DATA_BLOCK "T-104_Write_TO_Centrifuge_DB"   // DB309
TITLE = Signal Exchange between R-201<->Reactor_Selector
{ S7_Optimized_Access := 'TRUE' }
VERSION : 0.1
   VAR
      Wait : Bool;
      Started : Bool;   // Start Sequence
      Ready : Bool;
      Stop : Bool;   // Stop Sequence
      Abort : Bool;   // Abort Sequence
      Complete : Bool;
      Release : Bool;
      PARA : Bool;
      Initialization : Bool;
      PM : Bool;
      Monitoring : Bool;
      PumpingOut : Bool;   // Transfer to Cooling Tank
      PumpsOff : Bool;
      Held : Bool;   // Held Sequence
   END_VAR
BEGIN
END_DATA_BLOCK

DATA_BLOCK "T-104_Read_FROM_Centrifuge_DB"   // DB324
TITLE = Signal Exchange between R-201<->Reactor_Selector
{ S7_Optimized_Access := 'TRUE' }
VERSION : 0.1
   VAR
      StartTank : Bool;
      ReqWater : Bool;
      StopReqWater : Bool;
      Transfering : Bool;
      Pumps_OFF : Bool;
      Abort : Bool;
      Abort_Done : Bool;
      "Transfer_To_T-103_Done" : Bool;
      Idle : Bool;
   END_VAR
BEGIN
END_DATA_BLOCK

// folder: State MACHINE/1)Tanks/Tank T-104 (Water System)/T-104 <---> R-201

DATA_BLOCK "T-104_Write_TO_R-201_DB"   // DB287
TITLE = Signal Exchange between R-201<->Reactor_Selector
{ S7_Optimized_Access := 'TRUE' }
VERSION : 0.1
   VAR
      TankStarted : Bool;   // Start Sequence
      TankReady : Bool;
      Stop : Bool;   // Stop Sequence
      Abort : Bool;   // Abort Sequence
      PumpingOut : Bool;   // Transfer to Cooling Tank
      PumpsOff : Bool;
      Held : Bool;   // Held Sequence
   END_VAR
BEGIN
END_DATA_BLOCK

DATA_BLOCK "T-104_Read_FROM_R-201_DB"   // DB288
TITLE = Signal Exchange between R-201<->Reactor_Selector
{ S7_Optimized_Access := 'TRUE' }
VERSION : 0.1
   VAR
      StartTank : Bool;
      ReqWaterToWash : Bool;
      StopReqWaterToWash : Bool;
      ReqWater : Bool;
      StopReqWaterToPouring : Bool;
      Release : Bool;
      Abort : Bool;
      Abort_Done : Bool;
      Idle : Bool;
   END_VAR
BEGIN
END_DATA_BLOCK

// folder: State MACHINE/1)Tanks/Tank T-104 (Water System)/T-104 <---> R-202

DATA_BLOCK "T-104_Write_TO_R-202_DB"   // DB317
TITLE = Signal Exchange between R-201<->Reactor_Selector
{ S7_Optimized_Access := 'TRUE' }
VERSION : 0.1
   VAR
      TankStarted : Bool;   // Start Sequence
      TankReady : Bool;
      Stop : Bool;   // Stop Sequence
      Abort : Bool;   // Abort Sequence
      PumpingOut : Bool;   // Transfer to Cooling Tank
      PumpsOff : Bool;
      Held : Bool;   // Held Sequence
   END_VAR
BEGIN
END_DATA_BLOCK

DATA_BLOCK "T-104_Read_FROM_R-202_DB"   // DB318
TITLE = Signal Exchange between R-201<->Reactor_Selector
{ S7_Optimized_Access := 'TRUE' }
VERSION : 0.1
   VAR
      StartTank : Bool;
      ReqWaterToWash : Bool;
      StopReqWaterToWash : Bool;
      ReqWater : Bool;
      StopReqWaterToPouring : Bool;
      Release : Bool;
      Abort : Bool;
      Abort_Done : Bool;
      Idle : Bool;
   END_VAR
BEGIN
END_DATA_BLOCK

// folder: State MACHINE/1)Tanks/Tank T-104 (Water System)/T-104 <---> T-101

DATA_BLOCK "T-104_Read_FROM_T-101_DB"   // DB334
TITLE = Signal Exchange between R-201<->Reactor_Selector
{ S7_Optimized_Access := 'TRUE' }
VERSION : 0.1
   VAR
      StartTank : Bool;
      ReqWaterToWash : Bool;
      StopReqWaterToWash : Bool;
      ReqWaterToMix : Bool;
      StopReqWaterToMix : Bool;
      Release : Bool;
      Abort : Bool;
      Abort_Done : Bool;
      Idle : Bool;
   END_VAR
BEGIN
END_DATA_BLOCK

DATA_BLOCK "T-104_Write_TO_T-101_DB"   // DB341
TITLE = Signal Exchange between R-201<->Reactor_Selector
{ S7_Optimized_Access := 'TRUE' }
VERSION : 0.1
   VAR
      Wait : Bool;
      Started : Bool;   // Start Sequence
      Ready : Bool;
      Stop : Bool;   // Stop Sequence
      Abort : Bool;   // Abort Sequence
      Complete : Bool;
      Release : Bool;
      PARA : Bool;
      Initialization : Bool;
      PM : Bool;
      Monitoring : Bool;
      PumpingOut : Bool;   // Transfer to Cooling Tank
      PumpsOff : Bool;
      Held : Bool;   // Held Sequence
   END_VAR
BEGIN
END_DATA_BLOCK

// folder: State MACHINE/1)Tanks/Tank T-104 (Water System)/T-104 <---> T-102

DATA_BLOCK "T-104_Read_FROM_T-102_DB"   // DB337
TITLE = Signal Exchange between R-201<->Reactor_Selector
{ S7_Optimized_Access := 'TRUE' }
VERSION : 0.1
   VAR
      StartTank : Bool;
      ReqWaterToWash : Bool;
      StopReqWaterToWash : Bool;
      ReqWaterToMix : Bool;
      StopReqWaterToMix : Bool;
      Release : Bool;
      Abort : Bool;
      Abort_Done : Bool;
      Idle : Bool;
   END_VAR
BEGIN
END_DATA_BLOCK

DATA_BLOCK "T-104_Write_TO_T-102_DB"   // DB338
TITLE = Signal Exchange between R-201<->Reactor_Selector
{ S7_Optimized_Access := 'TRUE' }
VERSION : 0.1
   VAR
      Wait : Bool;
      Started : Bool;   // Start Sequence
      Ready : Bool;
      Stop : Bool;   // Stop Sequence
      Abort : Bool;   // Abort Sequence
      Complete : Bool;
      Release : Bool;
      PARA : Bool;
      Initialization : Bool;
      PM : Bool;
      Monitoring : Bool;
      PumpingOut : Bool;   // Transfer to Cooling Tank
      PumpsOff : Bool;
      Held : Bool;   // Held Sequence
   END_VAR
BEGIN
END_DATA_BLOCK

// folder: State MACHINE/2)Reactors/Reactor R-201

DATA_BLOCK "R-201_DB"   // DB268
{ S7_Optimized_Access := 'TRUE' }
VERSION : 0.1
   VAR
      Cmds : "UnitCmds";
      Status : Struct
         Initializing : Bool;
         Ready : Bool;
         Running : Bool;
         PouringRunning : Bool;
         TankWashRunning : Bool;
         TubeWashRunning : Bool;
         Aborting : Bool;
         Status : Int;   // 1=Idle, 2=Running, 3=Stopping, 4=Held, 5=Holding
         "Step" : Int;
         State : Int;
      END_STRUCT;
      OS : Struct
         bit : Array[0..15] of Bool;   // One Shot Bit
      END_STRUCT;
      Equipments : Struct
         Valves : Struct
            "XV-2013" : "Cmd";
            "XV-2011" : "Cmd";
            "XV-2021" : "Cmd";
            "XV-1043" : "Cmd";
            "FV-2011" : "Cmd";
            "FV-2021" : "Cmd";
         END_STRUCT;
         Pumps : Struct
            "P-201A" : "Cmd";
            "P-201B" : "Cmd";
         END_STRUCT;
         VFD : Struct
            "VFD-2011" : "Cmd";
         END_STRUCT;
      END_STRUCT;
      "Time" : Struct
         "Pre-Mix" : Time;   // Pre-Mix Time Displaying in the HMI
         pH_Delay : Time;   // pH Stabilize Time Displaying in the HMI
         Reaction : Time;   // Reaction Time Displaying in the HMI
         Wash : Time;   // Wash Time Displaying in the HMI
         Tube : Time;   // Tube Wash Time Displaying in the HMI
      END_STRUCT;
      PmpSel : Struct
         "P-201AB" : Int := 1;
      END_STRUCT;
   END_VAR
BEGIN
END_DATA_BLOCK

DATA_BLOCK "R-201_SEQ_DB"   // DB271
{ S7_Optimized_Access := 'TRUE' }
VERSION : 0.1
// stored: InstanceOfName R-201_SEQ
"R-201_SEQ"
BEGIN
END_DATA_BLOCK

DATA_BLOCK "R-201_Recipe"   // DB303
{ S7_Optimized_Access := 'TRUE' }
VERSION : 0.1
   VAR RETAIN
      Water : Real;   // Amount of Water to the Reactor before Pouring
   END_VAR
   VAR
      Temperature : Real := 80.0;   // Reactor Temperature
      MinLevelMixerOn : Real := 19.0;   // Minimum Level to Run the Mixer
      X_Flow : Real := 1.0;   // T-101(X) Flow to Transfer to Reactor
      Y_Flow : Real := 1.5;   // T-102(Y) Flow to Transfer to Reactor with pH Stability.
      X_Volume : Real;   // T-101(X) Volume to Transfer to Reactor
      LastWaterVolume : Real := 120.0;
      pH : Real := 8.0;   // pH Setpoint to the Reactor
      "Pre-Mix_Time" : Time := T#5m;   // Pre-Mix Time to the T-101 and T-102 before Transfer to Reactor
      pHStab_Time : Time := T#1m;   // Time to Stabilize the pH
      Reaction_Time : Time := T#22.5h;   // Reaction Time
   END_VAR
BEGIN
END_DATA_BLOCK

DATA_BLOCK "R-201_Aux_DB"   // DB354
{ S7_Optimized_Access := 'TRUE' }
VERSION : 0.1
   VAR
      "Real" : Struct
         "HFC-201" : Struct   // Heater
            SP : Real;
            Min : Real;   // Heater Minimum Temperature
            Max : Real;   // Heater Maximum Temperature
         END_STRUCT;
         PH : Struct   // pH Controller
            SP : Real;   // pH Set Point
            Min : Real;
            Max : Real;
         END_STRUCT;
         "FIC-2011" : Struct   // Fow Controller
            SP : Real := 1.0;   // Flow Setpoint
         END_STRUCT;
         "FIC-2021" : Struct
            SP : Real := 1.5;   // Flow Setpoint
         END_STRUCT;
         "T-101" : Struct
            TOTVolSP : Real;
         END_STRUCT;
         "LT-2011" : Struct
            Min : Real;
         END_STRUCT;
         "FT-1043" : Struct
            SP : Real;
         END_STRUCT;
         "VFD-R201" : Struct
            Start : Bool;
            Stop : Bool;
         END_STRUCT;
      END_STRUCT;
      "Timer" : Struct
         PreMix : IEC_TIMER;   // Timer Premix
         StabpH : IEC_TIMER;
         Reactor : IEC_TIMER;
         FlushOut : IEC_TIMER;
         MixToClean : IEC_TIMER;
         "XV-2013" : IEC_TIMER;
         "XV-2011" : IEC_TIMER;
         "XV-2021" : IEC_TIMER;
         "XV-1043" : IEC_TIMER;
         "FV-2011" : IEC_TIMER;
         "FV-2021" : IEC_TIMER;
      END_STRUCT;
      "Bool" : Struct
         PreMixT_En : Bool;   // Pre-Mix Timer Enable
         PreMixT_Reset : Bool;
         StabpHTEnStep : Bool;   // Stabilizer Timer Enable
         StabpHTEn : Bool;
         StabpHTEn_Reset : Bool;
         ReactorTEn : Bool;   // Enable Reacting time for the Reactor
         ReactorT_Reset : Bool;
         FlushOutTEn : Bool;
         MixToCleanTEn : Bool;   // Enable Timer to clean the reactor after Reacting
         MixToCleanT_Reset : Bool;
         TOff : Bool;   // Turning Off Valves
         Transitions : Struct
            TankEmpty : Bool;
         END_STRUCT;
      END_STRUCT;
      Constants : Struct
         CmdDelay : Time := T#2s;
      END_STRUCT;
   END_VAR
BEGIN
   "Timer".FlushOut.PT := T#5S;
   "Timer".PreMix.PT := T#5m;
   "Timer".StabpH.PT := T#1m;
   "Timer".MixToClean.PT := T#10M;
   "Timer".Reactor.PT := T#22.5h;
END_DATA_BLOCK

DATA_BLOCK "R-201_HMI_DB"   // DB358
{ S7_Optimized_Access := 'TRUE' }
VERSION : 0.1
   VAR
      FromHMI : "FromHMI";
      ToHMI : "ToHMI";
   END_VAR
BEGIN
END_DATA_BLOCK

// folder: State MACHINE/2)Reactors/Reactor R-201/Control R-201

DATA_BLOCK "R-201_Control_SEQ_DB"   // DB283
{ S7_Optimized_Access := 'TRUE' }
VERSION : 0.1
// stored: InstanceOfName R-201_Control
"R-201_Control"
BEGIN
END_DATA_BLOCK

DATA_BLOCK "R-201_Control_DB"   // DB300
{ S7_Optimized_Access := 'TRUE' }
VERSION : 0.1
   VAR
      FromHMI : Struct
         Start : Bool;
         Initialize : Bool;
         TankWash : Bool;
         TubeWash : Bool;
         Abort : Bool;
      END_STRUCT;
      Cmds : Struct
         Start : Bool;
         Initialize : Bool;
         TankWash : Bool;
         TubeWash : Bool;
         TransferToCoolingTank : Bool;
         Abort : Bool;
      END_STRUCT;
      Status : Struct
         Starting : Bool;
         Aborting : Bool;
      END_STRUCT;
      OS : Struct
         bit : Array[0..15] of Bool;   // One Shot Bit
      END_STRUCT;
   END_VAR
BEGIN
END_DATA_BLOCK

// folder: State MACHINE/2)Reactors/Reactor R-201/Control R-201/Control <---> R-201

DATA_BLOCK "Control_Write_TO_R-201_DB"   // DB277
TITLE = Signal Exchange between R-201<->Reactor_Selector
{ S7_Optimized_Access := 'TRUE' }
VERSION : 0.1
   VAR
      Wait : Bool;
      Start : Bool;   // Start Sequence
      Stop : Bool;   // Stop Sequence
      Abort : Bool;   // Abort Sequence
      Complete : Bool;
      Release : Bool;
      PARA : Bool;
      Initialization : Bool;
      PM : Bool;
      Running : Bool;
      WaitForTransfer : Bool;
      "Transfer_To_T-103" : Bool;   // Transfer to Cooling Tank
      TankWash : Bool;
      TubingWash : Bool;
      Held : Bool;   // Held Sequence
   END_VAR
BEGIN
END_DATA_BLOCK

DATA_BLOCK "Control_Read_FROM_R-201_DB"   // DB280
TITLE = Signal Exchange between R-201<->Reactor_Selector
{ S7_Optimized_Access := 'TRUE' }
VERSION : 0.1
   VAR
      ReactorStarted : Bool;
      Initialization_Done : Bool;
      Reacting_Done : Bool;
      Abort_Done : Bool;
      "Transfer_To_T-103_Done" : Bool;
      TankWash_done : Bool;
      TubeWash_Done : Bool;
      Idle : Bool;
   END_VAR
BEGIN
END_DATA_BLOCK

// folder: State MACHINE/2)Reactors/Reactor R-201/R-201 <---> Control

DATA_BLOCK "R-201_Write_TO_Control_DB"   // DB281
TITLE = Signal Exchange between R-201<->Reactor_Selector
{ S7_Optimized_Access := 'TRUE' }
VERSION : 0.1
   VAR
      ReactorStarted : Bool;
      Initialization_Done : Bool;
      Reacting_Done : Bool;
      Abort_Done : Bool;
      "Transfer_To_T-103_Done" : Bool;
      TankWash_done : Bool;
      TubeWash_Done : Bool;
      Idle : Bool;
   END_VAR
BEGIN
END_DATA_BLOCK

DATA_BLOCK "R-201_Read_FROM_Control_DB"   // DB282
TITLE = Signal Exchange between R-201<->Reactor_Selector
{ S7_Optimized_Access := 'TRUE' }
VERSION : 0.1
   VAR
      Wait : Bool;
      Start : Bool;   // Start Sequence
      Stop : Bool;   // Stop Sequence
      Abort : Bool;   // Abort Sequence
      Complete : Bool;
      Release : Bool;
      PARA : Bool;
      Initialization : Bool;
      PM : Bool;
      Running : Bool;
      WaitForTransfer : Bool;
      "Transfer_To_T-103" : Bool;   // Transfer to Cooling Tank
      TankWash : Bool;
      TubingWash : Bool;
      Held : Bool;   // Held Sequence
   END_VAR
BEGIN
END_DATA_BLOCK

// folder: State MACHINE/2)Reactors/Reactor R-201/R-201 <---> T-101

DATA_BLOCK "R-201_Read_FROM_T-101_DB"   // DB307
TITLE = Signal Exchange between R-201<->Reactor_Selector
{ S7_Optimized_Access := 'TRUE' }
VERSION : 0.1
   VAR
      TankStarted : Bool;   // Start Sequence
      Recirculating : Bool;
      PupmsOFF : Bool;   // Stop Sequence
      Abort : Bool;   // Abort Sequence
      RouteOpened : Bool;   // Transfer to Cooling Tank
      Idle : Bool;   // Held Sequence
   END_VAR
BEGIN
END_DATA_BLOCK

DATA_BLOCK "R-201_Write_TO_T-101_DB"   // DB327
TITLE = Signal Exchange between R-201<->Reactor_Selector
{ S7_Optimized_Access := 'TRUE' }
VERSION : 0.1
   VAR
      StartPouring : Bool;
      ReactorStarted : Bool;
      OpenRoute : Bool;
      RouteOpened : Bool;
      Transfering : Bool;
      FillingDone : Bool;
      Abort : Bool;
      Abort_Done : Bool;
      ReleaseTank : Bool;
      Idle : Bool;
   END_VAR
BEGIN
END_DATA_BLOCK

// folder: State MACHINE/2)Reactors/Reactor R-201/R-201 <---> T-102

DATA_BLOCK "R-201_Read_FROM_T-102_DB"   // DB316
TITLE = Signal Exchange between R-201<->Reactor_Selector
{ S7_Optimized_Access := 'TRUE' }
VERSION : 0.1
   VAR
      TankStarted : Bool;   // Start Sequence
      Recirculating : Bool;
      PupmsOFF : Bool;   // Stop Sequence
      Abort : Bool;   // Abort Sequence
      RouteOpened : Bool;   // Transfer to Cooling Tank
      Idle : Bool;   // Held Sequence
   END_VAR
BEGIN
END_DATA_BLOCK

DATA_BLOCK "R-201_Write_TO_T-102_DB"   // DB319
TITLE = Signal Exchange between R-201<->Reactor_Selector
{ S7_Optimized_Access := 'TRUE' }
VERSION : 0.1
   VAR
      StartPouring : Bool;
      ReactorStarted : Bool;
      OpenRoute : Bool;
      RouteOpened : Bool;
      Transfering : Bool;
      FillingDone : Bool;
      Abort : Bool;
      Abort_Done : Bool;
      ReleaseTank : Bool;
      Idle : Bool;
   END_VAR
BEGIN
END_DATA_BLOCK

// folder: State MACHINE/2)Reactors/Reactor R-201/R-201 <---> T-103 (CoolingTank)

DATA_BLOCK "R-201_Write_TO_T-103_DB"   // DB293
TITLE = Signal Exchange between R-201<->Reactor_Selector
{ S7_Optimized_Access := 'TRUE' }
VERSION : 0.1
   VAR
      StartTank : Bool;
      OpenRoute : Bool;
      Transfering : Bool;
      TubWash_Done : Bool;
      Abort : Bool;
      Abort_Done : Bool;
      "Transfer_To_T-103_Done" : Bool;
      Idle : Bool;
   END_VAR
BEGIN
END_DATA_BLOCK

DATA_BLOCK "R-201_Read_FROM_T-103_DB"   // DB296
TITLE = Signal Exchange between R-201<->Reactor_Selector
{ S7_Optimized_Access := 'TRUE' }
VERSION : 0.1
   VAR
      TankStarted : Bool;   // Start Sequence
      Stop : Bool;   // Stop Sequence
      Abort : Bool;   // Abort Sequence
      RouteOpened : Bool;   // Transfer to Cooling Tank
      Release : Bool;
      Held : Bool;   // Held Sequence
   END_VAR
BEGIN
END_DATA_BLOCK

// folder: State MACHINE/2)Reactors/Reactor R-201/R-201 <---> T-104 (WaterSystem)

DATA_BLOCK "R-201_Write_TO_T-104_DB"   // DB294
TITLE = Signal Exchange between R-201<->Reactor_Selector
{ S7_Optimized_Access := 'TRUE' }
VERSION : 0.1
   VAR
      StartTank : Bool;
      ReqWaterToWash : Bool;
      StopReqWaterToWash : Bool;
      ReqWater : Bool;
      StopReqWaterToPouring : Bool;
      Release : Bool;
      Abort : Bool;
      Abort_Done : Bool;
      Idle : Bool;
   END_VAR
BEGIN
END_DATA_BLOCK

DATA_BLOCK "R-201_Read_FROM_T-104_DB"   // DB295
TITLE = Signal Exchange between R-201<->Reactor_Selector
{ S7_Optimized_Access := 'TRUE' }
VERSION : 0.1
   VAR
      Wait : Bool;
      TankStarted : Bool;   // Start Sequence
      Ready : Bool;
      Stop : Bool;   // Stop Sequence
      Abort : Bool;   // Abort Sequence
      PumpingOut : Bool;   // Transfer to Cooling Tank
      PumpsOff : Bool;
      Held : Bool;   // Held Sequence
   END_VAR
BEGIN
END_DATA_BLOCK

// folder: State MACHINE/2)Reactors/Reactor R-202

DATA_BLOCK "R-202_DB"   // DB269
{ S7_Optimized_Access := 'TRUE' }
VERSION : 0.1
   VAR
      FromHMI : Struct
         Start : Bool;
         Initialize : Bool;
         TankWash : Bool;
         TubeWash : Bool;
         TransferToCoolingTank : Bool;
         Abort : Bool;
      END_STRUCT;
      Cmds : "UnitCmds";
      Status : Struct
         Initializing : Bool;
         Ready : Bool;
         Running : Bool;
         PouringRunning : Bool;
         TankWashRunning : Bool;
         TubeWashRunning : Bool;
         Aborting : Bool;
         Status : Int;   // 1=Idle, 2=Running, 3=Stopping, 4=Held, 5=Holding
         "Step" : Int;
         State : Int;
      END_STRUCT;
      OS : Struct
         bit : Array[0..15] of Bool;   // One Shot Bit
      END_STRUCT;
      Equipments : Struct
         Valves : Struct
            "XV-2023" : "Cmd";
            "XV-2012" : "Cmd";
            "XV-2022" : "Cmd";
            "XV-1044" : "Cmd";
            "FV-2012" : "Cmd";
            "FV-2022" : "Cmd";
         END_STRUCT;
         Pumps : Struct
            "P-202A" : "Cmd";
            "P-202B" : "Cmd";
         END_STRUCT;
         VFD : Struct
            "VFD-2021" : "Cmd";
         END_STRUCT;
      END_STRUCT;
      "Time" : Struct
         "Pre-Mix" : Time;   // Pre-Mix Time Displaying in the HMI
         PH_Delay : Time;   // pH Stabilize Time Displaying in the HMI
         Reaction : Time;   // Reaction Time Displaying in the HMI
         Wash : Time;   // Wash Time Displaying in the HMI
         Tube : Time;   // Tube Wash Time Displaying in the HMI
      END_STRUCT;
      PmpSel : Struct
         "P-202AB" : Int := 1;
      END_STRUCT;
   END_VAR
BEGIN
END_DATA_BLOCK

DATA_BLOCK "R-202_SEQ_DB"   // DB286
{ S7_Optimized_Access := 'TRUE' }
VERSION : 0.1
// stored: InstanceOfName R-202_SEQ
"R-202_SEQ"
BEGIN
END_DATA_BLOCK

DATA_BLOCK "R-202_Recipe"   // DB304
{ S7_Optimized_Access := 'TRUE' }
VERSION : 0.1
   VAR RETAIN
      Water : Real;   // Amount of Water to the Reactor before Pouring
   END_VAR
   VAR
      Temperature : Real := 80.0;   // Reactor Temperature
      MinLevelMixerOn : Real := 19.0;   // Minimum Level to Run the Mixer
      X_Flow : Real := 1.0;   // T-101(X) Flow to Transfer to Reactor
      Y_Flow : Real := 1.5;   // T-102(Y) Flow to Transfer to Reactor with pH Stability.
      X_Volume : Real;   // T-101(X) Volume to Transfer to Reactor
      LastWaterVolume : Real := 120.0;
      pH : Real := 8.0;   // pH Setpoint to the Reactor
      "Pre-Mix_Time" : Time := T#5m;   // Pre-Mix Time to the T-101 and T-102 before Transfer to Reactor
      pHStab_Time : Time := T#1m;   // Time to Stabilize the pH
      Reaction_Time : Time := T#22.5h;   // Reaction Time
   END_VAR
BEGIN
END_DATA_BLOCK

DATA_BLOCK "R-202_Aux_DB"   // DB365
{ S7_Optimized_Access := 'TRUE' }
VERSION : 0.1
   VAR
      "Real" : Struct
         "HFC-201" : Struct   // Heater
            SP : Real;
            Min : Real;   // Heater Minimum Temperature
            Max : Real;   // Heater Maximum Temperature
         END_STRUCT;
         PH : Struct   // pH Controller
            SP : Real;   // pH Set Point
            Min : Real;
            Max : Real;
         END_STRUCT;
         "FIC-2012" : Struct   // Fow Controller
            SP : Real;   // Flow Setpoint
         END_STRUCT;
         "FIC-2022" : Struct
            SP : Real := 1.0;   // Flow Setpoint
         END_STRUCT;
         "T-101" : Struct
            TOTVolSP : Real;
         END_STRUCT;
         "LT-2021" : Struct
            Min : Real;
         END_STRUCT;
         "FT-1044" : Struct
            SP : Real;
         END_STRUCT;
         "VFD-R202" : Struct
            Start : Bool;
            Stop : Bool;
         END_STRUCT;
      END_STRUCT;
      "Timer" : Struct
         PreMix : IEC_TIMER;   // Timer Premix
         StabpH : IEC_TIMER;
         Reactor : IEC_TIMER;
         FlushOut : IEC_TIMER;
         MixToClean : IEC_TIMER;
         "XV-2023" : IEC_TIMER;
         "XV-2012" : IEC_TIMER;
         "XV-2022" : IEC_TIMER;
         "XV-1044" : IEC_TIMER;
         "FV-2012" : IEC_TIMER;
         "FV-2022" : IEC_TIMER;
      END_STRUCT;
      "Bool" : Struct
         PreMixT_En : Bool;   // Pre-Mix Timer Enable
         PreMixT_Reset : Bool;
         StabpHTEnStep : Bool;   // Stabilizer Timer Enable
         StabpHTEn : Bool;   // Stabilizer Timer Enable
         StabpHTEn_Reset : Bool;
         ReactorTEn : Bool;   // Enable Reacting time for the Reactor
         ReactorT_Reset : Bool;
         FlushOutTEn : Bool;
         MixToCleanTEn : Bool;   // Enable Timer to clean the reactor after Reacting
         MixToCleanT_Reset : Bool;
         TOff : Bool;   // Turning Off Valves
         Transitions : Struct
            TankEmpty : Bool;
         END_STRUCT;
      END_STRUCT;
      Constants : Struct
         CmdDelay : Time := T#2s;
      END_STRUCT;
   END_VAR
BEGIN
   "Timer".FlushOut.PT := T#5S;
   "Timer".PreMix.PT := T#5m;
   "Timer".StabpH.PT := T#1m;
   "Timer".MixToClean.PT := T#10M;
   "Timer".Reactor.PT := T#21.5h;
END_DATA_BLOCK

DATA_BLOCK "R-202_HMI_DB"   // DB367
{ S7_Optimized_Access := 'TRUE' }
VERSION : 0.1
   VAR
      FromHMI : "FromHMI";
      ToHMI : "ToHMI";
   END_VAR
BEGIN
END_DATA_BLOCK

// folder: State MACHINE/2)Reactors/Reactor R-202/Control R-202

DATA_BLOCK "R-202_Control_SEQ_DB"   // DB290
{ S7_Optimized_Access := 'TRUE' }
VERSION : 0.1
// stored: InstanceOfName R-202_Control
"R-202_Control"
BEGIN
END_DATA_BLOCK

DATA_BLOCK "R-202_Control_DB"   // DB344
{ S7_Optimized_Access := 'TRUE' }
VERSION : 0.1
   VAR
      FromHMI : Struct
         Start : Bool;
         Initialize : Bool;
         TankWash : Bool;
         TubeWash : Bool;
         Abort : Bool;
      END_STRUCT;
      Cmds : Struct
         Start : Bool;
         Initialize : Bool;
         TankWash : Bool;
         TubeWash : Bool;
         Abort : Bool;
      END_STRUCT;
      Status : Struct
         Starting : Bool;
         Aborting : Bool;
      END_STRUCT;
      OS : Struct
         bit : Array[0..15] of Bool;   // One Shot Bit
      END_STRUCT;
   END_VAR
BEGIN
END_DATA_BLOCK

// folder: State MACHINE/2)Reactors/Reactor R-202/Control R-202/Control <---> R-202

DATA_BLOCK "Control_Write_TO_R-202_DB"   // DB270
TITLE = Signal Exchange between R-201<->Reactor_Selector
{ S7_Optimized_Access := 'TRUE' }
VERSION : 0.1
   VAR
      Wait : Bool;
      Start : Bool;   // Start Sequence
      Stop : Bool;   // Stop Sequence
      Abort : Bool;   // Abort Sequence
      Complete : Bool;
      Release : Bool;
      PARA : Bool;
      Initialization : Bool;
      PM : Bool;
      Running : Bool;
      "Transfer_To_T-103" : Bool;   // Transfer to Cooling Tank
      TankWash : Bool;
      TubingWash : Bool;
      Held : Bool;   // Held Sequence
   END_VAR
BEGIN
END_DATA_BLOCK

DATA_BLOCK "Control_Read_FROM_R-202_DB"   // DB273
TITLE = Signal Exchange between R-201<->Reactor_Selector
{ S7_Optimized_Access := 'TRUE' }
VERSION : 0.1
   VAR
      ReactorStarted : Bool;
      Initialization_Done : Bool;
      Reacting_Done : Bool;
      Abort_Done : Bool;
      "Transfer_To_T-103_Done" : Bool;
      TankWash_done : Bool;
      TubeWash_Done : Bool;
      Idle : Bool;
   END_VAR
BEGIN
END_DATA_BLOCK

// folder: State MACHINE/2)Reactors/Reactor R-202/R-202 <---> Control

DATA_BLOCK "R-202_Write_TO_Control_DB"   // DB285
TITLE = Signal Exchange between R-201<->Reactor_Selector
{ S7_Optimized_Access := 'TRUE' }
VERSION : 0.1
   VAR
      ReactorStarted : Bool;
      Initialization_Done : Bool;
      Reacting_Done : Bool;
      Abort_Done : Bool;
      "Transfer_To_T-103_Done" : Bool;
      TankWash_done : Bool;
      TubeWash_Done : Bool;
      Idle : Bool;
   END_VAR
BEGIN
END_DATA_BLOCK

DATA_BLOCK "R-202_Read_FROM_Control_DB"   // DB289
TITLE = Signal Exchange between R-201<->Reactor_Selector
{ S7_Optimized_Access := 'TRUE' }
VERSION : 0.1
   VAR
      Wait : Bool;
      Start : Bool;   // Start Sequence
      Stop : Bool;   // Stop Sequence
      Abort : Bool;   // Abort Sequence
      Complete : Bool;
      Release : Bool;
      PARA : Bool;
      Initialization : Bool;
      PM : Bool;
      Running : Bool;
      "Transfer_To_T-103" : Bool;   // Transfer to Cooling Tank
      TankWash : Bool;
      TubingWash : Bool;
      Held : Bool;   // Held Sequence
   END_VAR
BEGIN
END_DATA_BLOCK

// folder: State MACHINE/2)Reactors/Reactor R-202/R-202 <---> T-101

DATA_BLOCK "R-202_Read_FROM_T-101_DB"   // DB312
TITLE = Signal Exchange between R-201<->Reactor_Selector
{ S7_Optimized_Access := 'TRUE' }
VERSION : 0.1
   VAR
      TankStarted : Bool;   // Start Sequence
      Recirculating : Bool;
      PupmsOFF : Bool;   // Stop Sequence
      Abort : Bool;   // Abort Sequence
      RouteOpened : Bool;   // Transfer to Cooling Tank
      Idle : Bool;   // Held Sequence
   END_VAR
BEGIN
END_DATA_BLOCK

DATA_BLOCK "R-202_Write_TO_T-101_DB"   // DB329
TITLE = Signal Exchange between R-201<->Reactor_Selector
{ S7_Optimized_Access := 'TRUE' }
VERSION : 0.1
   VAR
      StartPouring : Bool;
      ReactorStarted : Bool;
      OpenRoute : Bool;
      RouteOpened : Bool;
      Transfering : Bool;
      FillingDone : Bool;
      Abort : Bool;
      Abort_Done : Bool;
      ReleaseTank : Bool;
      Idle : Bool;
   END_VAR
BEGIN
END_DATA_BLOCK

// folder: State MACHINE/2)Reactors/Reactor R-202/R-202 <---> T-102

DATA_BLOCK "R-202_Read_FROM_T-102_DB"   // DB313
TITLE = Signal Exchange between R-201<->Reactor_Selector
{ S7_Optimized_Access := 'TRUE' }
VERSION : 0.1
   VAR
      TankStarted : Bool;   // Start Sequence
      Recirculating : Bool;
      PupmsOFF : Bool;   // Stop Sequence
      Abort : Bool;   // Abort Sequence
      RouteOpened : Bool;   // Transfer to Cooling Tank
      Idle : Bool;   // Held Sequence
   END_VAR
BEGIN
END_DATA_BLOCK

DATA_BLOCK "R-202_Write_TO_T-102_DB"   // DB330
TITLE = Signal Exchange between R-201<->Reactor_Selector
{ S7_Optimized_Access := 'TRUE' }
VERSION : 0.1
   VAR
      StartPouring : Bool;
      ReactorStarted : Bool;
      OpenRoute : Bool;
      RouteOpened : Bool;
      Transfering : Bool;
      FillingDone : Bool;
      Abort : Bool;
      Abort_Done : Bool;
      ReleaseTank : Bool;
      Idle : Bool;
   END_VAR
BEGIN
END_DATA_BLOCK

// folder: State MACHINE/2)Reactors/Reactor R-202/R-202 <---> T-103 (CoolingTank)

DATA_BLOCK "R-202_Write_TO_T-103_DB"   // DB332
TITLE = Signal Exchange between R-201<->Reactor_Selector
{ S7_Optimized_Access := 'TRUE' }
VERSION : 0.1
   VAR
      StartTank : Bool;
      OpenRoute : Bool;
      Transfering : Bool;
      TubWash_Done : Bool;
      Abort : Bool;
      Abort_Done : Bool;
      "Transfer_To_T-103_Done" : Bool;
      Idle : Bool;
   END_VAR
BEGIN
END_DATA_BLOCK

DATA_BLOCK "R-202_Read_FROM_T-103_DB"   // DB343
TITLE = Signal Exchange between R-201<->Reactor_Selector
{ S7_Optimized_Access := 'TRUE' }
VERSION : 0.1
   VAR
      TankStarted : Bool;   // Start Sequence
      Stop : Bool;   // Stop Sequence
      Abort : Bool;   // Abort Sequence
      RouteOpened : Bool;   // Transfer to Cooling Tank
      Release : Bool;
      Held : Bool;   // Held Sequence
   END_VAR
BEGIN
END_DATA_BLOCK

// folder: State MACHINE/2)Reactors/Reactor R-202/R-202 <---> T-104 (WaterSystem)

DATA_BLOCK "R-202_Write_TO_T-104_DB"   // DB335
TITLE = Signal Exchange between R-201<->Reactor_Selector
{ S7_Optimized_Access := 'TRUE' }
VERSION : 0.1
   VAR
      StartTank : Bool;
      ReqWaterToWash : Bool;
      StopReqWaterToWash : Bool;
      ReqWater : Bool;
      StopReqWaterToPouring : Bool;
      Release : Bool;
      Abort : Bool;
      Abort_Done : Bool;
      Idle : Bool;
   END_VAR
BEGIN
END_DATA_BLOCK

DATA_BLOCK "R-202_Read_FROM_T-104_DB"   // DB339
TITLE = Signal Exchange between R-201<->Reactor_Selector
{ S7_Optimized_Access := 'TRUE' }
VERSION : 0.1
   VAR
      Wait : Bool;
      TankStarted : Bool;   // Start Sequence
      Ready : Bool;
      Stop : Bool;   // Stop Sequence
      Abort : Bool;   // Abort Sequence
      PumpingOut : Bool;   // Transfer to Cooling Tank
      PumpsOff : Bool;
      Held : Bool;   // Held Sequence
   END_VAR
BEGIN
END_DATA_BLOCK

// folder: State MACHINE/3)Centrifuge

DATA_BLOCK "Centrifuge_DB"   // DB266
{ S7_Optimized_Access := 'TRUE' }
VERSION : 0.1
   VAR
      Transitions : Struct
         "T-103_Empty" : Bool;
         WaterDone : Bool;
         InitialsDone : Bool;
         ReadytoRun : Bool;
         BasketFull : Bool;
      END_STRUCT;
      Timers : Struct
         BucketTimerDelay : IEC_TIMER;
      END_STRUCT;
      Cmds : "UnitCmds";
      Status : Struct
         Initializing : Bool;
         Ready : Bool;
         Running : Bool;
         PouringRunning : Bool;
         TankWashRunning : Bool;
         TubeWashRunning : Bool;
         Aborting : Bool;
         Status : Int;   // 1=Idle, 2=Running, 3=Stopping, 4=Held, 5=Holding
         "Step" : Int;
         State : Int;
      END_STRUCT;
      OS : Struct
         bit : Array[0..15] of Bool;   // One Shot Bit
      END_STRUCT;
      Equipments : Struct
         Valves : Struct
            "XV-1045" : "Cmd";
            "XV-3013" : "Cmd";
            "XV-3012" : "Cmd";
            "XV-3011" : "Cmd";
            "FV-3011" : "Cmd";
         END_STRUCT;
         Pumps : Struct
            "P-301A" : "Cmd";
            "P-301B" : "Cmd";
         END_STRUCT;
         VFD : Struct
            "C-3011" : "Centrifuge";
         END_STRUCT;
      END_STRUCT;
      "Time" : Struct
         DrySpin : Time;
      END_STRUCT;
      PmpSel : Struct   // PumpSelection
         "P-301AB" : Int := 1;   // 1=P-301A, 2=P-301B
      END_STRUCT;
   END_VAR
BEGIN
END_DATA_BLOCK

DATA_BLOCK "Centrifuge_SEQ_DB"   // DB299
{ S7_Optimized_Access := 'TRUE' }
VERSION : 0.1
// stored: InstanceOfName Centrifuge_SEQ
"Centrifuge_SEQ"
BEGIN
END_DATA_BLOCK

DATA_BLOCK "Centrifuge_Aux_DB"   // DB356
{ S7_Optimized_Access := 'TRUE' }
VERSION : 0.1
   VAR
      "Real" : Struct
         "FIC-3011" : Struct
            SP : Real := 10.0;
         END_STRUCT;
         "VFD-3011" : Struct
            SP : Real := 50.0;
         END_STRUCT;
         "FT-3011" : Struct
            SP : Real := 280.0;
         END_STRUCT;
         DryTime : Struct
            SP : Time := T#10M;
         END_STRUCT;
      END_STRUCT;
      "Int" : Struct
         CentrifugeSpeedFbk : Int;
      END_STRUCT;
      "Timer" : Struct
         "XV-1045" : IEC_TIMER;
         "XV-3013" : IEC_TIMER;
         "XV-3012" : IEC_TIMER;
         "XV-3011" : IEC_TIMER;
         "FV-3011" : IEC_TIMER;
         WaitForBucket : IEC_TIMER;
         DryingWetCake : IEC_TIMER;
         DrySpinDnDelay : IEC_TIMER;   // Dry Spin Done Delay to Finish
      END_STRUCT;
      "Bool" : Struct
         TOff : Bool;   // Turning Off Valves
         WaitForBucketEn : Bool;   // Wait for get some Level in the Bucket before Start Pumps
         DryingWetCakeEn : Bool;   // Run the Pumps after Turn off the Water to dry the wet cake
         DryingWetCake_Reset : Bool;
         DrySpinDnDelay_Enab : Bool;
         Centrifuge : Struct
            Status : Struct
               MotorRunning : Bool;
               VibrationFault : Bool;
               ESTOP : Bool;
               SystemFault : Bool;
               BasketFull : Bool;
               CoverLocked : Bool;
               FeelerRetracted : Bool;
               FeelerEngaged : Bool;
            END_STRUCT;
            Command : Struct
               Start : Bool;
               Stop : Bool;
               ESTOP : Bool := TRUE;   // ESTOP to Centrifuge, 1=OK
               RetFeelerAndReset : Bool;
               FeelerEngage : Bool;
            END_STRUCT;
         END_STRUCT;
      END_STRUCT;
      Constants : Struct
         CmdDelay : Time := T#2s;
      END_STRUCT;
   END_VAR
BEGIN
   "Timer".DryingWetCake.PT := t#30m;
   "Timer".DrySpinDnDelay.PT := T#30s;
END_DATA_BLOCK

DATA_BLOCK "Centrifuge_HMI_DB"   // DB363
{ S7_Optimized_Access := 'TRUE' }
VERSION : 0.1
   VAR
      FromHMI : "FromHMI";
      ToHMI : "ToHMI";
      FromHMI_Aux : Struct
         Start : Bool;   // Start Centrifuge
         Stop : Bool;   // Stop Centrifuge
         FeelerRetReset : Bool;   // Feeler Retrac and Reset
         FeelerEngage : Bool;   // Feeler Engage
      END_STRUCT;
   END_VAR
BEGIN
END_DATA_BLOCK

// folder: State MACHINE/3)Centrifuge/Centrifuge <---> T-103

DATA_BLOCK "Centrifuge_Write_TO_T-103_DB"   // DB310
TITLE = Signal Exchange between R-201<->Reactor_Selector
{ S7_Optimized_Access := 'TRUE' }
VERSION : 0.1
   VAR
      RequestProduct : Bool;   // Request Product
      OpenRoute : Bool;
      RouteOpened : Bool;   // Abort Sequence
      "T-103_Empty" : Bool;   // T-103 Tank empty
      BasketFull : Bool;   // Basket Full Signal
      FeelerRet : Bool;   // Feeler Retracted
      CloseRoute : Bool;
      Release : Bool;
   END_VAR
BEGIN
END_DATA_BLOCK

DATA_BLOCK "Centrifuge_Read_FROM_T-103_DB"   // DB320
TITLE = Signal Exchange between R-201<->Reactor_Selector
{ S7_Optimized_Access := 'TRUE' }
VERSION : 0.1
   VAR
      ReadyToTransfer : Bool;
      Done : Bool;
      RouteOpened : Bool;
      Transfering : Bool;
      Pumps_OFF : Bool;
      Abort : Bool;
      Abort_Done : Bool;
      "Transfer_To_T-103_Done" : Bool;
      Idle : Bool;
   END_VAR
BEGIN
END_DATA_BLOCK

// folder: State MACHINE/3)Centrifuge/Centrifuge <---> T-104

DATA_BLOCK "Centrifuge_Write_TO_T-104_DB"   // DB315
TITLE = Signal Exchange between R-201<->Reactor_Selector
{ S7_Optimized_Access := 'TRUE' }
VERSION : 0.1
   VAR
      StartTank : Bool;   // Start Sequence
      ReqWater : Bool;
      StopReqWater : Bool;
      Abort : Bool;   // Abort Sequence
      Complete : Bool;
      Release : Bool;
      PARA : Bool;
      Initialization : Bool;
      PM : Bool;
      Monitoring : Bool;
      RouteOpened : Bool;   // Transfer to Cooling Tank
      Held : Bool;   // Held Sequence
   END_VAR
BEGIN
END_DATA_BLOCK

DATA_BLOCK "Centrifuge_Read_FROM_T-104_DB"   // DB323
TITLE = Signal Exchange between R-201<->Reactor_Selector
{ S7_Optimized_Access := 'TRUE' }
VERSION : 0.1
   VAR
      Wait : Bool;
      Started : Bool;   // Start Sequence
      Ready : Bool;
      Stop : Bool;   // Stop Sequence
      Abort : Bool;   // Abort Sequence
      Complete : Bool;
      Release : Bool;
      PARA : Bool;
      Initialization : Bool;
      PM : Bool;
      Monitoring : Bool;
      PumpingOut : Bool;   // Transfer to Cooling Tank
      PumpsOff : Bool;
      Held : Bool;   // Held Sequence
   END_VAR
BEGIN
END_DATA_BLOCK

// folder: State MACHINE/4)Calcination

DATA_BLOCK "R401_TempMon_DB"   // DB20
{ S7_Optimized_Access := 'TRUE' }
AUTHOR : JLopez
VERSION : 0.1
// stored: InstanceOfName AI Monitor
"AI Monitor"
BEGIN
END_DATA_BLOCK

DATA_BLOCK "Calcination_DB"   // DB91
{ S7_Optimized_Access := 'TRUE' }
VERSION : 0.1
   VAR
      Alarms : Struct
         Communication : Struct
            Fault : Bool;
         END_STRUCT;
      END_STRUCT;
      Shutdowns : Struct
         "1 Activated" : Bool;
         "2 Activated" : Bool;
      END_STRUCT;
      MonBlockData : Struct
         Input : Struct
            AvgSP : Real;   // Average SP Furnace Temperature
            "Min Range" : Real;   // Minimum Furnace Temperature Range
            "Max Range" : Real;   // Maximun Furnace Temperature Range
            MinAvgValue : Real := 0.0;   // Min Average Hysteresis Range
            MaxAvgValue : Real := 0.0;   // Max Average Hysteresis Range
            EnableDeviationMon : Bool;
            AlarmDeviation : Real := 0.0;
            MaxDeviation : Real := 0.0;   // Maximun deviation Allows
            MaxAboveTemp : Real := 50.0;
         END_STRUCT;
         Output : Struct
            Avg : Real;   // Average Value
            AvgReached : Bool;   // Average Reached (Actual Average >=Avg-Minimum Average and <=Avg+Maximum Average
            AvgAlarm : Bool;
            ReadyToProcess : Bool;   // Conditions meet(Average,Range,Deviation) and ready to operate
            DeviationAlarm : Bool;
            DeviationFault : Bool;   // Deviation Fault Activated
            MaxAboveTempFault : Bool;   // Max Above Temperature Fault Activated
         END_STRUCT;
      END_STRUCT;
   END_VAR
   VAR RETAIN
      CalcinationTimeSp : Time := T#2h;
   END_VAR
   VAR
      CicleCnt : Int;   // Cicle Counter
      ControlSEQ : Struct
         AbortSeq : Bool;
         AbortDone : Bool;
         OS : Array[0..31] of Bool;
         TestBits : Array[0..31] of Bool;
      END_STRUCT;
   END_VAR
BEGIN
   // ControlSEQ.OS[0] : Abort SEQUENCE
END_DATA_BLOCK

DATA_BLOCK "R-401_AIMon_DB"   // DB241
{ S7_Optimized_Access := 'TRUE' }
AUTHOR : JLopez
VERSION : 0.1
// stored: InstanceOfName AI Monitor_v2
"AI Monitor_v2"
BEGIN
END_DATA_BLOCK

DATA_BLOCK "Calcination_HMI_DB"   // DB366
{ S7_Optimized_Access := 'TRUE' }
VERSION : 0.1
   VAR
      FromHMI : Struct
         Start : Bool;   // Start Sequence
         Stop : Bool;   // Stop Sequence
         Pause : Bool;
         Initialize : Bool;   // Initialize Sequence
         TankWash : Bool;   // Tank Wash Procedure
         TubeWash : Bool;   // Line Wash Procedure
         TransferToCoolingTank : Bool;   // Transfer to Cooling Tank (T-103)
      END_STRUCT;
      ToHMI : Struct
         EnStopButton : Bool;   // Enable HMI Stop Button
         EnStartButton : Bool;   // Enable HMI Start Button
         EnRestartButton : Bool;
         EnPauseButton : Bool;
         EnOpeRequest : Bool;   // Enable HMI Operator Request Button
         EnEditorButton : Bool;   // Enable HMI Editor Burron Button
      END_STRUCT;
   END_VAR
BEGIN
END_DATA_BLOCK

// folder: State MACHINE/4)Calcination/Reactor R-401

DATA_BLOCK "R-401_Recipe"   // DB92
{ S7_Optimized_Access := 'TRUE' }
VERSION : 0.1
   VAR
      Temperature : Struct
         SP1 : Real := 300.0;   // R-401 Set Point 1 to Temperature Controller
         SP2 : Real := 400.0;   // R-401 Set Point 2 to Temperature Controller
         SP3 : Real := 750.0;   // R-401 Set Point 3 to Temperature Controller
         NormalShutdown : Real := 30.0;
         "Slow Shutdown" : Real := 28.0;   // R-401 Slow Shutdown Temperature
         RampRate : Struct
            SP1 : Int := 3;   // Heat Up Ramp 1 (degress/min)
            SP2 : Int := 3;   // Heat Up Ramp 2 (degress/min)
            SP3 : Int := 3;   // Heat Up Ramp 3 (degress/min)
            "Cold Down" : Int := 10;   // Cold Down Ramp (degress/min)
         END_STRUCT;
         Dwell : Struct
            SP1 : Int := 180;
            SP2 : Int := 180;
            SP3 : Int := 180;
         END_STRUCT;
      END_STRUCT;
      Pressure : Struct
         Air : Real := 16.2;   // R-401 Pressure
         N2 : Real := 16.2;
         Shutdown : Real := 0.0;   // R-401 Shutdown Pressure
      END_STRUCT;
      CalcinationTime : Struct
         SP1 : Time := T#1H;   // Calcination Time Setpoint
         SP2 : Time := T#1H;
         SP3 : Time := T#2H;
      END_STRUCT;
   END_VAR
BEGIN
END_DATA_BLOCK

DATA_BLOCK "R-401_SEQ_DB"   // DB377
{ S7_Optimized_Access := 'TRUE' }
AUTHOR : JL
VERSION : 0.1
// stored: InstanceOfName R-401_SEQ
"R-401_SEQ"
BEGIN
END_DATA_BLOCK

DATA_BLOCK "R-401_DB"   // DB378
{ S7_Optimized_Access := 'TRUE' }
VERSION : 0.1
   VAR
      Transitions : Struct
         "T-103_Empty" : Bool;
         WaterDone : Bool;
      END_STRUCT;
      Timers : Struct
         BucketTimerDelay : IEC_TIMER;
      END_STRUCT;
      Cmds : "UnitCmds";
      Status : Struct
         Initializing : Bool;
         Ready : Bool;
         Running : Bool;
         Spare1 : Bool;
         Spare2 : Bool;
         ShuttingDown : Bool;   // Controlled Shutting Down
         Aborting : Bool;
         Status : Int;   // 1=Idle, 2=Running, 3=Stopping, 4=Held, 5=Holding
         "Step" : Int;
         State : Int;
      END_STRUCT;
      OS : Struct
         bit : Array[0..15] of Bool;   // One Shot Bit
      END_STRUCT;
      Equipments : Struct
         Valves : Struct
            "FV-4011" : "Cmd";
            "FV-4012" : "Cmd";
            "TC-4011" : "Cmd";
         END_STRUCT;
         Pumps : Struct
            "P-301A" : "Cmd";
            "P-301B" : "Cmd";
         END_STRUCT;
         VFD : Struct
            "VFD-3011" : "Cmd_VFD";
         END_STRUCT;
      END_STRUCT;
      "Time" : Struct
         HoldTime : Time;
      END_STRUCT;
      PmpSel : Struct   // PumpSelection
         "P-301AB" : Int := 1;   // 1=P-301A, 2=P-301B
      END_STRUCT;
   END_VAR
BEGIN
END_DATA_BLOCK

DATA_BLOCK "R-401_Aux_DB"   // DB379
{ S7_Optimized_Access := 'TRUE' }
VERSION : 0.1
   VAR
      "Real" : Struct
         "TE-401" : Struct
            Temperature : Struct
               MinRange : Real := 50.0;
               MaxRange : Real := 50.0;
               MinAvgValue : Real := 1.0;
               MaxAvgValue : Real := 30.0;
               AlarmDeviation : Real := 25.0;
               MaxDeviation : Real := 50.0;
            END_STRUCT;
         END_STRUCT;
         "MFC-4011" : Struct
            Pressure : Struct
               Min : Real := 0.0;   // R-401 Shutdown Pressure
               Max : Real;
            END_STRUCT;
         END_STRUCT;
         "MFC-4012" : Struct
            Pressure : Struct
               Min : Real := 0.0;   // R-401 Shutdown Pressure
               Max : Real;
            END_STRUCT;
         END_STRUCT;
      END_STRUCT;
      "Timer" : Struct
         "FV-4011" : IEC_TIMER;
         "FV-4012" : IEC_TIMER;
         "TC-4011" : IEC_TIMER;
         HoldTime : Struct
            SP : Time := T#1h;   // Hold Time Setpoint
         END_STRUCT;
         HoldTimer : IEC_TIMER;
         CalcinationTime : Struct
            SP : Time := T#10m;   // Calcination Time Setpoint
         END_STRUCT;
         CalcinationTimer : IEC_TIMER;   // Calcination Timer
      END_STRUCT;
      "Bool" : Struct
         TOff : Bool;   // Turning Off Valves
         ShutdownAux : Bool;   // Shutdown Auxiliar bit
         CalcinationTimeEn : Bool;
         CalcinationTime_Reset : Bool;
         HoldTimeEn : Bool;
         HoldTime_Reset : Bool;
         Cond : Struct
            _001 : Bool;   // Cond: Average Temperature reached, Timer Done, Cotroller Reseted
            _002 : Bool;   // Temperature Setpoints Send and received
            _003 : Bool;   // Ramp Rate Setpoints Send and received
            _004 : Bool;   // Dwell Setpoints Send and received
            _005 : Bool;   // Setpoitns Sent
            _006 : Bool;   // Working SP Reached the SP A
            _007 : Bool;   // Working SP Reached the SP B
            _008 : Bool;   // Working SP Reached the SP C
            _009 : Bool;   // All Working SP are the same
         END_STRUCT;
      END_STRUCT;
      Constants : Struct
         CmdDelay : Time := T#2s;
      END_STRUCT;
   END_VAR
BEGIN
END_DATA_BLOCK

DATA_BLOCK "R-401_HMI_DB"   // DB380
{ S7_Optimized_Access := 'TRUE' }
VERSION : 0.1
   VAR
      FromHMI : "FromHMI";
      ToHMI : "ToHMI";
   END_VAR
BEGIN
END_DATA_BLOCK

// folder: State MACHINE/5)Passivate

DATA_BLOCK "Passivation_HMI_DB"   // DB368
{ S7_Optimized_Access := 'TRUE' }
VERSION : 0.1
   VAR
      FromHMI : Struct
         Start : Bool;   // Start Sequence
         Stop : Bool;   // Stop Sequence
         Pause : Bool;
         Initialize : Bool;   // Initialize Sequence
         TankWash : Bool;   // Tank Wash Procedure
         TubeWash : Bool;   // Line Wash Procedure
         TransferToCoolingTank : Bool;   // Transfer to Cooling Tank (T-103)
      END_STRUCT;
      ToHMI : Struct
         EnStopButton : Bool;   // Enable HMI Stop Button
         EnStartButton : Bool;   // Enable HMI Start Button
         EnRestartButton : Bool;
         EnPauseButton : Bool;
         EnOpeRequest : Bool;   // Enable HMI Operator Request Button
         EnEditorButton : Bool;   // Enable HMI Editor Burron Button
      END_STRUCT;
   END_VAR
BEGIN
END_DATA_BLOCK

DATA_BLOCK "Mon_R402_DB"   // DB413
{ S7_Optimized_Access := 'TRUE' }
AUTHOR : JLopez
VERSION : 0.1
// stored: InstanceOfName AI Monitor
"AI Monitor"
BEGIN
END_DATA_BLOCK

// folder: State MACHINE/5)Passivate/Reactor R-402

DATA_BLOCK "R-402_Recipe"   // DB387
{ S7_Optimized_Access := 'TRUE' }
VERSION : 0.1
   VAR
      Temperature : Struct
         SP1 : Real := 365.0;   // R-401 Set Point 1 to Temperature Controller
         SP2 : Real := 400.0;   // R-401 Set Point 2 to Temperature Controller
         SP3 : Real := 750.0;   // R-401 Set Point 3 to Temperature Controller
         NormalShutdown : Real := 30.0;
         "Slow Shutdown" : Real := 25.0;   // R-401 Slow Shutdown Temperature
         RampRate : Struct
            SP1 : Int := 10;   // Heat Up Ramp 1 (degress/min)
            SP2 : Int := 3;   // Heat Up Ramp 2 (degress/min)
            SP3 : Int := 3;   // Heat Up Ramp 3 (degress/min)
            "Cold Down" : Int := 10;   // Cold Down Ramp (degress/min)
         END_STRUCT;
      END_STRUCT;
      Reduction : Struct
         "N2 Pressure SP" : Real := 18.5;   // N2 Pressure Setpoint
         "H2 Flow SP" : Real := 1.0;   // H2 Flow Setpoint
         Shutdown : Real := 0.0;   // Shutdown Pressure
      END_STRUCT;
      Passivation : Struct
         "Air Pressure SP" : Real := 0.02;   // Air Pressure SP
         "H2 Flow SP" : Real;   // H2 Flow Setpoint
         Shutdown : Real := 0.0;   // Shutdown Pressure
      END_STRUCT;
      HoldTime : Struct
         SP1 : Time := T#2H;   // Time Setpoint 1
         SP2 : Time;   // Time Setpoint 2
         SP3 : Time;   // Time Setpoint 3
      END_STRUCT;
   END_VAR
BEGIN
END_DATA_BLOCK

DATA_BLOCK "R-402_DB"   // DB399
{ S7_Optimized_Access := 'TRUE' }
VERSION : 0.1
   VAR
      Transitions : Struct
         xxx : Bool;
      END_STRUCT;
      Timers : Struct
         xxx : IEC_TIMER;
      END_STRUCT;
      Cmds : "UnitCmds";
      Status : Struct
         Initializing : Bool;
         Ready : Bool;
         Running : Bool;
         Spare1 : Bool;
         Spare2 : Bool;
         ShuttingDown : Bool;   // Controlled Shutting Down
         Aborting : Bool;
         Status : Int;   // 1=Idle, 2=Running, 3=Stopping, 4=Held, 5=Holding
         "Step" : Int;
         State : Int;
      END_STRUCT;
      OS : Struct
         bit : Array[0..15] of Bool;   // One Shot Bit
      END_STRUCT;
      Equipments : Struct
         Valves : Struct
            "XV-4021" : "Cmd";
            "XV-4022" : "Cmd";
            "XV-4024" : "Cmd";
            "XV-4025" : "Cmd";
            "FV-4021" : "Cmd";
            "FV-4024" : "Cmd";
            "FV-4025" : "Cmd";
            "TC-402A" : "Cmd";
            "TC-402B" : "Cmd";
         END_STRUCT;
      END_STRUCT;
      "Time" : Struct
         HoldTime : Time;
      END_STRUCT;
      PmpSel : Struct   // PumpSelection
         xxx : Int := 1;   // 1=P-301A, 2=P-301B
      END_STRUCT;
   END_VAR
BEGIN
END_DATA_BLOCK

DATA_BLOCK "R-402_Aux_DB"   // DB400
{ S7_Optimized_Access := 'TRUE' }
VERSION : 0.1
   VAR
      "Real" : Struct
         "TE-402" : Struct
            Temperature : Struct
               MinRange : Real := 50.0;
               MaxRange : Real := 50.0;
               MinAvgValue : Real := 5.0;
               MaxAvgValue : Real := 5.0;
               AlarmDeviation : Real := 25.0;
               MaxDeviation : Real := 50.0;
            END_STRUCT;
         END_STRUCT;
         "MFC-4025" : Struct
            Pressure : Struct
               Min : Real := 0.0;   // R-401 Pressure
               Max : Real := 0.0;   // R-401 Shutdown Pressure
            END_STRUCT;
         END_STRUCT;
      END_STRUCT;
      "Timer" : Struct
         "XV-4021" : IEC_TIMER;
         "XV-4022" : IEC_TIMER;
         "XV-4024" : IEC_TIMER;
         "XV-4025" : IEC_TIMER;
         "FV-4021" : IEC_TIMER;
         "FV-4024" : IEC_TIMER;
         "FV-4025" : IEC_TIMER;
         "TC-402" : IEC_TIMER;
         HoldTime : Struct
            SP : Time := T#10M;   // Hold Time Setpoint
         END_STRUCT;
         HoldTimer : IEC_TIMER;
         CalcinationTime : Struct
            SP : Time := T#10M;   // Calcination Time Setpoint
         END_STRUCT;
         CalcinationTimer : IEC_TIMER;   // Calcination Timer
         Alarms : Struct
            MFC_Cmms1 : IEC_TIMER;
            MFC_Cmms2 : IEC_TIMER;
            "TC-4011A_Cmms1" : IEC_TIMER;
            "TC-4011A_Cmms2" : IEC_TIMER;
            "TC-4011B_Cmms1" : IEC_TIMER;
            "TC-4011B_Cmms2" : IEC_TIMER;
            "TC-4011C_Cmms1" : IEC_TIMER;
            "TC-4011C_Cmms2" : IEC_TIMER;
         END_STRUCT;
      END_STRUCT;
      "Bool" : Struct
         TOff : Bool;   // Turning Off Valves
         ShutdownAux : Bool;   // Shutdown Auxiliar bit
         CalcinationTimeEn : Bool;
         CalcinationTime_Reset : Bool;
         HoldTimeEn : Bool;
         HoldTime_Reset : Bool;
         Cond : Struct
            _001 : Bool;   // Cond: Average Temperature reached, Timer Done, Cotroller Reseted
            _002 : Bool;   // Temperature Setpoints Send and received
            _003 : Bool;   // Ramp Rate Setpoints Send and received
            _004 : Bool;   // Dwell Setpoints Send and received
            _005 : Bool;   // Setpoitns Sent
            _006 : Bool;   // Working SP Reached the SP A
            _007 : Bool;   // Working SP Reached the SP B
            _008 : Bool;   // Working SP Reached the SP C
            _009 : Bool;   // All Working SP are the same
         END_STRUCT;
         EurothermStatus : Struct
            "4011A_Connected" : Bool;   // 1=Controllers Conected, 0=No connection
            "4011B_Connected" : Bool;   // 1=Controllers Conected, 0=No connection
            "4011C_Connected" : Bool;   // 1=Controllers Conected, 0=No connection
         END_STRUCT;
      END_STRUCT;
      Constants : Struct
         CmdDelay : Time := T#2s;
      END_STRUCT;
   END_VAR
BEGIN
END_DATA_BLOCK

DATA_BLOCK "R-402_HMI_DB"   // DB401
{ S7_Optimized_Access := 'TRUE' }
VERSION : 0.1
   VAR
      FromHMI : "FromHMI";
      ToHMI : "ToHMI";
   END_VAR
BEGIN
END_DATA_BLOCK

DATA_BLOCK "R-402_SEQ_DB"   // DB414
{ S7_Optimized_Access := 'TRUE' }
AUTHOR : JL
VERSION : 0.1
// stored: InstanceOfName R-402_SEQ
"R-402_SEQ"
BEGIN
END_DATA_BLOCK

// folder: System blocks/Program resources

DATA_BLOCK "StartCentrifuge_Pulse"   // DB164
{ S7_Optimized_Access := 'TRUE' }
AUTHOR : Simatic
FAMILY : IEC
NAME : IEC_TMR
VERSION : 1.0
// stored: InstanceOfName IEC_TIMER
"IEC_TIMER"
BEGIN
END_DATA_BLOCK

DATA_BLOCK "StopCentrifuge_Pulse"   // DB167
{ S7_Optimized_Access := 'TRUE' }
AUTHOR : Simatic
FAMILY : IEC
NAME : IEC_TMR
VERSION : 1.0
// stored: InstanceOfName IEC_TIMER
"IEC_TIMER"
BEGIN
END_DATA_BLOCK

DATA_BLOCK "CentrifugeFeelerRetractAndReset"   // DB169
{ S7_Optimized_Access := 'TRUE' }
AUTHOR : Simatic
FAMILY : IEC
NAME : IEC_TMR
VERSION : 1.0
// stored: InstanceOfName IEC_TIMER
"IEC_TIMER"
BEGIN
END_DATA_BLOCK

DATA_BLOCK "CentrifugeFeelerEngage"   // DB173
{ S7_Optimized_Access := 'TRUE' }
AUTHOR : Simatic
FAMILY : IEC
NAME : IEC_TMR
VERSION : 1.0
// stored: InstanceOfName IEC_TIMER
"IEC_TIMER"
BEGIN
END_DATA_BLOCK

DATA_BLOCK "T-103_Empty_Condition_C"   // DB298
{ S7_Optimized_Access := 'TRUE' }
AUTHOR : Simatic
FAMILY : IEC
NAME : IEC_TMR
VERSION : 1.0
// stored: InstanceOfName IEC_TIMER
"IEC_TIMER"
BEGIN
END_DATA_BLOCK

// folder: Timers

DATA_BLOCK "interlock_Timers"   // DB244
{ S7_Optimized_Access := 'TRUE' }